FUNCTION_BLOCK "LKinCtrl_MC_MovePath"   // FB35000, SCL
TITLE = LKinCtrl_MovePath
{ S7_Optimized_Access := 'TRUE' }
AUTHOR : tech.team.motioncontrol@siemens.com
FAMILY : LKinCtrl
VERSION : 3.0
// Core function block of LKinCtrl library:
// executes path motion provided by PathData command list
   VAR_INPUT
      execute : Bool;   // rising edge starts action once
      stop : Bool;   // abort path motion
      interrupt : Bool;   // interrupt path motion
      reset : Bool;   // reset FB / acknowledge errors
      sequenceMode : Int;   // activate sequence mode (0) / single step mode (1)
      pathTransition : DInt;   // initial transition configuration for new path motion (1: use bufferMode and transitionParameter)
      bufferMode : DInt := 1;   // inital bufferMode for new path motion
      transitionParameter : Array[1..5] of LReal;   // initial transitionParameter for new path motion
      configuration : "LKinCtrl_typeConfiguration";   // configuration structure
   END_VAR
   VAR_OUTPUT
      done : Bool;   // TRUE: Commanded functionality has been completed successfully
      busy : Bool;   // TRUE: FB is not finished and new output values can be expected
      active : Bool;   // FB in control of axesGroup / kinematic in motion
      commandAborted : Bool;   // TRUE: Commanded functionality has been aborted by another command
      error : Bool;   // TRUE: An error occurred during the execution of the FB
      status : Word;   // status of the FB
      diagnostics : "LKinCtrl_typeMovePathDiagnostics";   // diagnostics information of FB
      activePathData : String["LKINCTRL_LENGTH_OF_PATHDATA_NAME"];   // name of actual PathData
      activeCmdNo : DInt := 0;   // number of actual PathData set
      remainingDistanceActCmd : LReal;   // remaining distance of actual PathData set
      readyForNextPath : Bool := true;   // TRUE: Next PathData can be triggered
   END_VAR
   VAR_IN_OUT
      axesGroup : TO_Kinematics;   // reference to the axesGroup
      pathData : Variant;   // reference to the PathData
      flags : Array[0.."LKINCTRL_NO_OF_LAST_SETFLAG"] of Bool;   // boolean defined by setFlags in PathCommand
      valueFlags : Array[0.."LKINCTRL_NO_OF_LAST_VALUEFLAG"] of LReal;   // value defined by valueFlags in PathCommand
   END_VAR
   VAR
      statExecuteOld : Bool;   // old value of 'execute' input for edge detection
      statStopOld : Bool;   // old value of 'stop' input for edge detection
      statInterruptOld : Bool;   // old value of 'interrupt' input for edge detection
      statResetOld : Bool;   // old value of 'reset' input for edge detection
      statDone : Bool;   // static value for output 'done'
      statBusy : Bool;   // static value for output 'busy'
      statCommandAborted : Bool;   // static value for output 'commandAborted'
      statError : Bool;   // static value for output 'error'
      statErrorID : Word;   // flagWord for FB output: errorID
      statStatus : Word := 16#7000;   // static value for output 'status'
      statSubfunctionStatus : Word;   // status or return value of called FBs, FCs and system blocks
      statStateExecution : DInt := 0;   // state in the state machine of the FB
      statStatePreBuffering : DInt := 0;   // state in the state machine of the FB
      statDebugState : Bool;   // static variable to debug IF state machine if needed
      statEmptyDiagnostics : "LKinCtrl_typeMovePathDiagnostics";   // empty diagnostics information (for initialization purposes only)
      instLKinCtrl_MC_ExecuteKinMotionCmd : "LKinCtrl_MC_ExecuteKinMotionCmd";
      instLKinCtrl_PreBuffer : "LKinCtrl_PreBuffer";
      statPathDataPreBuffered : "LKinCtrl_typePathData_PreBuf";   // preBuffered PathData elements (internal buffer of path motion commands)
      statPathDataElementPreBuffered : "LKinCtrl_typePathDataElement_PreBuf";   // PathData element to be executed by FB_ExecutePathMotion
      statFlagsBuffer : Struct   // buffer to store flag information for past and actual commands
         writeBufferElement : Int := 1;   // pointer on entry to be written
         bufferElement : Array[1.."LKINCTRL_NO_OF_SETFLAGS_BUFFER_ELEMENTS"] of Struct   // flag information for one specific command (see cmdId)
            pathDataName : String["LKINCTRL_LENGTH_OF_PATHDATA_NAME"];   // PathData name of specific command
            pathDataIdentifier : DInt;   // PathData identifier counter of specific command
            cmdId : DInt;   // cmdId of command in PathData
            isIntermediateCmd : Bool;   // TRUE: command is intermediate command
            setFlags : Array[1.."LKINCTRL_NO_OF_CMD_SETFLAGS"] of "LKinCtrl_typeSetFlagElement_Bool";   // setFlags structure equal to PathData command entry
            valueFlags : Array[1.."LKINCTRL_NO_OF_CMD_VALUEFLAGS"] of "LKinCtrl_typeSetFlagElement_LReal";   // setFlags structure equal to PathData command entry
         END_STRUCT;
      END_STRUCT;
      statLastCmdIdPathdata : DInt;   // static value to store last detected cmd in PathData
      statPathDataPreBufferAddPointerOld : Int;   // old value of 'addPointer' in PathDataPreBuffer
      statReadyForNextPath : Bool := true;   // static value for output 'readyForNextPath'
      statStoreInterruptStateExecution : DInt;   // static store variable for state machine status on interrupt
      statExecutionWaitSingleStep : Bool;   // static bit to wait for execution due to sequenceMode
      statExecutionWaitTimerRunning : Bool;   // static bit to wait for execution due to wait time running
      statWaitMain : Bool;   // static bit to wait for execution due to wait flags
      statWaitValueMain : Bool;   // static bit to wait for execution due to wait value flags
      statPreBufferCmdCtr : Int;   // static counter to run FB LKinCtrl_PreBuffer multiple times
      statWaitFlags : Struct   // static struct to store wait flag information
         waitCtr : Int;   // counter for number of wait flags in one command
         waitFlag : Array[1.."LKINCTRL_NO_OF_CMD_SETFLAGS"] of Int;   // flag number as identifier for flag active as wait flag
      END_STRUCT;
      statWaitValueFlags : Struct   // static struct to store wait valueFlag information
         waitCtr : Int;   // counter for number of wait flags in one command
         waitFlag : Array[1.."LKINCTRL_NO_OF_CMD_VALUEFLAGS"] of Int;   // flag number as identifier for flag active as wait valueFlag
      END_STRUCT;
      statPreBufferedPathDataNameOld : String["LKINCTRL_LENGTH_OF_PATHDATA_NAME"];   // static to store old PathDataName in PathDataPreBuffered
      statPathDataIdentifier : USInt;   // static to identify PathDatas independent of given name
      statPreBufferedCmdIdOld : DInt;   // static to store old cmdId value from PathDataPreBuffered
      statSetFlagsBufferWriteBufferElement_old : Int;   // static to store old setFlagsBuffer write element pointer value
      statExecuterWasDone : Bool;   // static to store done output of executer in case of wait flags at end of path
      statWrittenActiveCmdNo : DInt;   // static to store the last written active command number
      statInterruptedAtStart : Bool;   // static to store if interrupt was executed at start of path
      statInitPos : Array[1..4] of LReal;   // static to store the initial position of the TCP
      statOCSFrames : Array[1..3] of "LKinCtrl_typeFrame";   // static to store the OCS frames from TO_Kinematics
      instLKinCtrl_SetFlagCtrl : "LKinCtrl_SetFlagCtrl";
      instLKinCtrl_ValueFlagCtrl : "LKinCtrl_ValueFlagCtrl";
   END_VAR
   VAR_TEMP
      tempExecute : Bool;   // Temporary value for input 'execute'
      tempStop : Bool;   // Temporary value for input 'stop'
      tempInterrupt : Bool;   // Temporary value for input 'interrupt'
      tempReset : Bool;   // Temporary value for input 'stop'
      tempSequenceMode : Int;   // Temporary value for input 'sequenceMode'
      tempEmptyPathDataElementPreBuffered : "LKinCtrl_typePathDataElement_PreBuf";   // Temporary value for empty pre buffer element
      tempCmdCtr : Int;   // Temporary command counter
      tempFlagsBufferElementCtr : Int;   // Temporary flag buffer counter
      tempPreBufferCallCtr : Int;   // Temporary flag buffer call counter
      tempFlagCmdCounter : Int;   // Temporary flag command counter
      tempFlagResetCmdCounter : Int;   // Temporary flag reset counter
   END_VAR
   VAR CONSTANT
      EX_NO_PROCESSING : Int := 0;   // state machine constant
      EX_RESETTING : Int := 5;   // state machine constant
      EX_INTERRUPT_AT_START : Int := 10;   // state machine constant
      EX_GET_CMD : Int := 30;   // state machine constant
      EX_TRIGGERING_CMD : Int := 50;   // state machine constant
      EX_TRIGGERED_CMD : Int := 55;   // state machine constant
      EX_INTERRUPTING : Int := 70;   // state machine constant
      EX_INTERRUPTED : Int := 75;   // state machine constant
      EX_CONTINUEING : Int := 77;   // state machine constant
      EX_CONTINUED : Int := 78;   // state machine constant
      EX_STOPPING : Int := 80;   // state machine constant
      EX_STOPPED_STATE : Int := 85;   // state machine constant
      EX_ERROR_STATE : Int := 90;   // state machine constant
      EX_ALL_TRIGGERED : Int := 100;   // state machine constant
      PB_NO_PROCESSING : Int := 0;   // state machine constant
      PB_ENABLED : Int := 10;   // state machine constant
      PB_OFF_COMP : Int := 15;   // state machine constant
      PB_DISABLED : Int := 20;   // state machine constant
      STATUS_EXECUTION_FINISHED : Word := 16#0000;   // status execution finished without errors
      STATUS_NO_CALL : Word := 16#7000;   // status no job being currently processed
      STATUS_FIRST_CALL : Word := 16#7001;   // status first call after incoming new job (rising edge 'execute')
      STATUS_SUBSEQUENT_CALL : Word := 16#7002;   // status subsequent call during active processing without further details
      STATUS_FB_RESETTING : Word := 16#7010;   // status FB resetting
      STATUS_WAITING_FOR_PREBUFFERED_CMD : Word := 16#7070;   // status waiting for new command in PathData_Prebuffered
      STATUS_PREBUFFERED_FULL : Word := 16#7071;   // status internal cmd buffer filled completely
      STATUS_CMD_LIN_ACTIVE : Word := 16#7301;   // status linear motion command active at axesgroup
      STATUS_CMD_CIRC_ACTIVE : Word := 16#7302;   // status circular motion command active at axesgroup
      STATUS_PATHMOTION_INTERRUPTED : Word := 16#7303;   // status path motion interrupted
      STATUS_PATHMOTION_STOPPING : Word := 16#7304;   // status path motion stopping
      STATUS_READYFORNEXTPATH : Word := 16#7305;   // status FB ready for next path execution
      STATUS_PATHMOTION_RUNNING : Word := 16#7306;   // status path motion running
      STATUS_EXECUTION_WAITING : Word := 16#7307;   // status path execution waiting due to wait flag, wait time or single step mode
      STATUS_CMD_MOVE_DIRECT_ACTIVE : Word := 16#7308;   // status move direct motion command active at axesgroup
      STATUS_STOP_DUE_TO_ERROR : Word := 16#7309;   // status kinematics is stopped due to an error in FB Executer
      STATUS_COMMAND_ABORTED : Word := 16#7FFF;   // status commanded functionality has been aborted by another command
      ERR_UNDEFINED_STATE : Word := 16#8600;   // error due to an undefined state in state machine
      ERR_EXECUTE_KINMOTIONCMD : Word := 16#8201;   // error due to error in FB LKinCtrl_ExecuteKinMotionCmd
      ERR_WRONG_SEQUENCEMODE : Word := 16#8203;   // error due to invalid sequenceMode on input
      ERR_PATHDATA_PARAMETERS : Word := 16#8204;   // error due to malconfiguration in motion command parameters
      ERR_OFFSET_CALCULATION : Word := 16#8205;   // error due to calculation error in offset compensation
      ERR_ERROR_STILL_PENDING : Word := 16#8207;   // error due to previous not acknowledged error (reset MovePath to acknowledge)
      ERR_SET_FLAG_CONTROL : Word := 16#8208;   // error due to error in set flag control FB
      ERR_VALUE_FLAG_CONTROL : Word := 16#8209;   // error due to error in value flag control FB
      INTERRUPT_AT_START : Bool := FALSE;   // interrupt at start of new path to preload commands
      NO_OF_COMMANDS_PRELOADING : USInt := 3;   // number of commands to be preloaded
   END_VAR
   // transitionParameter[1] := -1.0;
   // statFlagsBuffer.bufferElement[1].cmdId := 0;
   // statFlagsBuffer.bufferElement[1].pathDataName := '';
BEGIN
   //==========================================================================================
   // SIEMENS AG
   // (c)Copyright 2020 All Rights Reserved
   //------------------------------------------------------------------------------------------
   // Library: LKinCtrl
   // Tested with: S7-1517T-3 PN/DP
   // Engineering: TIA Portal V16
   // Restrictions: ---
   // Requirements: S7-1500T FW 2.8
   // Functionality: LKinCtrl_MC_MovePath
   // The FB is executing a sequence to drive a path defined by the user in form of a
   // command list of points and motion commands.
   // 
   // Support: tech.team.motioncontrol@siemens.com
   // Note: Parameter comments are only available in language 'English (United States)'
   //------------------------------------------------------------------------------------------
   // Change log table:
   // Version    Date          Expert in charge    Changes applied
   // 01.00.00   06.02.2018    JR                  First release version v1.0
   // 02.00.00   18.04.2019    JR / FR             V2.0
   // 02.01.00   28.05.2019    JR / FR             V2.1 for LKinLang
   // 02.02.00   28.01.2020    JR / FR             V2.2: Added valueFlags and flagOnlyCmd 
   // 02.02.01   07.02.2020    FR / DF             V2.2.1: Disable Prebuffer when MovePath is stopping/reseting/(done)
   // 02.02.02   12.02.2020    FR                  Fix for loops using wrong flag constant
   // 02.03.00   18.03.2020    FR                  Rework Flag FBs; Fix for interrupt/continue
   // 02.04.00   25.03.2020    FR                  Added preprocessing stop for LKinLang
   // 02.04.01   07.05.2020    FR                  Fix 360° circle with circMode 3
   // 02.04.02   16.07.2020    FR                  Several bugfixes
   // 03.00.00   04.08.2020    FR                  Added MoveDirect and ConveyorTracking; V16/FW2.8.2 required!
   // 03.00.01   06.08.2020    FR                  Bugfix
   // 03.00.02   19.10.2020    FR                  Updated ContourOffset; Updated FlagControl; Bugfixes
   // 03.00.03   23.11.2020    FR                  Updated ContourOffset; Fix in MC_ExecuteKinMotionCmd
   // 03.00.05   01.06.2021    FR                  Fixes in FlagCtrl FBs
   // 03.00.06   06.07.2021    FR                  Updated ContourOffset; Fix in MC_ExecuteKinMotionCmd; Fix in FlagCtrl FBs
   //===========================================================================================

   // Work with temporary value / create process image
   #tempExecute := #execute;
   #tempStop := #stop;
   #tempInterrupt := #interrupt;
   #tempReset := #reset;
   #tempSequenceMode := #sequenceMode;

   REGION TRIGGERING
       //===========================================================================================
       // check for sequenceMode to be activated
       IF #tempSequenceMode = 1 THEN
           // set execution wait bit to stop cmds from being executed (wait in EX_TRIGGERING_CMD)
           #statExecutionWaitSingleStep := TRUE;
           // check for incorrect sequenceMode to be selected
       ELSIF (#tempSequenceMode <> 0 AND #tempSequenceMode <> 1)
           // only check if execution is triggered
           AND #tempExecute = TRUE
       THEN
           // set status accordingly
           #statStatus := #ERR_WRONG_SEQUENCEMODE;
           // set execution state machine
           #statStateExecution := #EX_ERROR_STATE;
       END_IF;

       //===========================================================================================
       // check for rising edge of stop input
       IF (#tempStop = TRUE) AND (#statStopOld = FALSE)
       THEN
           // perform stop procedure
           #statStateExecution := #EX_STOPPING;
           // FR 08.04.2020: Set status and bits here to avoid return when status = STATUS_NO_CALL
           #statStatus := #STATUS_PATHMOTION_STOPPING;
           #statDone := FALSE;
           #statBusy := TRUE;
           #statCommandAborted := FALSE;
           #statError := FALSE;
           #statErrorID := 16#0;


           //===========================================================================================
           // check for rising edge of interrupt input
           // FR 17.03.2020: Added "statDone" to condition
           // FR 09.04.2020: Added stopping status to condition
       ELSIF (#tempInterrupt = TRUE) AND (#statInterruptOld = FALSE) AND (#statDone = FALSE)
           AND #statStatus <> #STATUS_PATHMOTION_STOPPING AND #statStatus <> #STATUS_COMMAND_ABORTED
       THEN
           // FR 11.03.2020: Only save state in some cases
           IF #statStateExecution < #EX_INTERRUPTING
               OR #statStateExecution > #EX_CONTINUED THEN
               // store states of interruption for later continue
               #statStoreInterruptStateExecution := #statStateExecution;
           END_IF;
           // perform interrupt procedure
           #statStateExecution := #EX_INTERRUPTING;
           //===========================================================================================
           // check for rising edge of reset input
       ELSIF (#tempReset = TRUE) AND (#statResetOld = FALSE)
           // interlock reset during execution
           AND (#statBusy = FALSE)
       THEN
           // perform reset procedure
           #statStateExecution := #EX_RESETTING;
           #statStatePreBuffering := #PB_NO_PROCESSING;
           // set status accordingly
           #statStatus := #STATUS_FB_RESETTING;
           //===========================================================================================
           // check for rising edge of execute input
       ELSIF (#tempExecute = TRUE) AND (#statExecuteOld = FALSE)
           AND (#stop = FALSE) AND (#interrupt = FALSE)
       THEN // First call; initialize FB
           #statDone := FALSE;
           #statCommandAborted := FALSE;
           #statError := FALSE;
           #statErrorID := 16#0;

           // ERROR on start
           //===========================================================================================
           // check for state machine to be in error state from previous (not acknowledged) error
           IF #statStateExecution = #EX_ERROR_STATE THEN
             // State machine - do not start cmd execution and wait in error state
             //------------------------------------------------------------------------------------------
             // no changes to PreBuffer state machine
             #statStateExecution := #EX_ERROR_STATE;
             #statStatePreBuffering := #PB_NO_PROCESSING;

             // check for error already detected before execute in this cycle (e.g. wrong sequenceMode / other faulty inputs)
             IF #statStatus = #ERR_WRONG_SEQUENCEMODE THEN
               // reset statBusy to avoid interlock of reset
               #statBusy := FALSE;
             ELSE
               // set status to set error bit
               #statStatus := #ERR_ERROR_STILL_PENDING;
             END_IF;


             // continue motion in SINGLESTEP mode
             //===========================================================================================
             // check for execution to be waiting for new rising edge
           ELSIF #statStateExecution = #EX_TRIGGERING_CMD
             AND #statExecutionWaitSingleStep = TRUE
           THEN
             // set FB state to busy
             #statBusy := TRUE;
             // reset execution wait bit stopping cmds from being executed (wait in EX_TRIGGERING_CMD)
             #statExecutionWaitSingleStep := FALSE;

             // CONTINUE after interrupt
             //===========================================================================================
             // check for path motion to be interrupted
           ELSIF #statStateExecution = #EX_INTERRUPTED THEN
             // State machine - continue path motion and sequence
             //------------------------------------------------------------------------------------------
             // no changes to PreBuffer state machine
             #statStateExecution := #EX_CONTINUEING;

             // no setting of FB state to busy necessary, interrupt does not reset busy

             // RETRIGGER during running path motion
             // ==========================================================================================
             // check for path motion to be running with all previous cmds executed
           ELSIF #statStateExecution = #EX_ALL_TRIGGERED
           THEN
             // set FB state to busy
             #statBusy := TRUE;

             // // reset last cmdId in PathData depending on type of attached PathData
             #statLastCmdIdPathdata := 0;

             // Reset bit to memorize done output of MC_ExecuteKinMotionCmd
             #statExecuterWasDone := FALSE;

             // state machines - reStart processing
             //------------------------------------------------------------------------------------------
             #statStatePreBuffering := #PB_ENABLED;
             #statStateExecution := #EX_GET_CMD;
             //------------------------------------------------------------------------------------------
             // initialize functionality: reset of variables, diagnostics, etc. (only at reTriggering)
             #statReadyForNextPath := FALSE;

             // set status - added JR 2019/04/16
             #statStatus := #STATUS_SUBSEQUENT_CALL;

             // START of path motion (initial)
             //===========================================================================================
             // check for path motion not to be running already
           ELSIF #axesGroup.StatusMotionQueue.NumberOfCommands = 0         // no commands in MotionQueue
             AND #axesGroup.StatusWord.%X12 = TRUE                       // TO Kinematics in constant velocity
             AND #axesGroup.StatusPath.Velocity = 0.0                    // TO Kinematics standing still
             AND (#axesGroup.StatusWord.%X6                              // no motion job in progress
             OR #axesGroup.StatusConveyor[1].TrackingState <> 0          // If kinematics is in tracking then done (.X6) is not set
             OR #axesGroup.StatusConveyor[2].TrackingState <> 0
             OR #axesGroup.StatusConveyor[3].TrackingState <> 0)
             AND #statStatus <> #STATUS_EXECUTION_WAITING                // Added FR 2019.03.28
           THEN
             //------------------------------------------------------------------------------------------
             // initialize functionality: reset of variables, diagnostics, etc. (only at first call, no reTriggering)
             #statStatus := #STATUS_FIRST_CALL;
             // set FB state to busy
             #statBusy := TRUE;
             #diagnostics := #statEmptyDiagnostics;
             #statSubfunctionStatus := 16#0;
             #statPathDataPreBuffered.addPointerRestarted := FALSE;

             // initialize buffer variables
             //------------------------------------------------------------------------------------------
             // delete PathDataPreBuffered
             FOR #tempCmdCtr := 1 TO "LKINCTRL_NO_OF_PATHDATA_PREBUFFER_ELEMENTS" DO
               #statPathDataPreBuffered.commands[#tempCmdCtr] := #tempEmptyPathDataElementPreBuffered;
             END_FOR;
             // reset PathDataPreBuffered retrievePointer
             #statPathDataPreBuffered.retrievePointer := 1;
             // initialize add pointer in PathData_PreBuffered
             #statPathDataPreBuffered.addPointer := 1;
             #statPathDataPreBuffered.pathDataName := '';
             // delete cmd stored for execution
             #statPathDataElementPreBuffered := #tempEmptyPathDataElementPreBuffered;
             // counter variable PreBuffer call cycles
             #statPreBufferCmdCtr := "LKINCTRL_NO_OF_START_EXECUTE_CMDS";

             // Reset bit to memorize done output of MC_ExecuteKinMotionCmd
             #statExecuterWasDone := FALSE;
             // reset storage static for old PathData identification value
             #statPathDataIdentifier := 0;

             // store actual position - in case of path starting with relative cmd for contour offset compensation
             //------------------------------------------------------------------------------------------
             #statInitPos[1] := #axesGroup.Tcp.x;
             #statInitPos[2] := #axesGroup.Tcp.y;
             #statInitPos[3] := #axesGroup.Tcp.z;
             #statInitPos[4] := #axesGroup.Tcp.a;

             // initialize flag handling variables
             //------------------------------------------------------------------------------------------
             // Reset waitFlags struct
             #statWaitFlags.waitCtr := 0;
             FOR #tempFlagResetCmdCounter := 1 TO "LKINCTRL_NO_OF_CMD_SETFLAGS" DO
               #statWaitFlags.waitFlag[#tempFlagResetCmdCounter] := -1;
             END_FOR;

             // Reset waitValueFlag struct
             #statWaitValueFlags.waitCtr := 0;
             FOR #tempFlagResetCmdCounter := 1 TO "LKINCTRL_NO_OF_CMD_VALUEFLAGS" DO
               #statWaitValueFlags.waitFlag[#tempFlagResetCmdCounter] := -1;
             END_FOR;

             // reset setFlagsBuffer variables
             #statFlagsBuffer.writeBufferElement := 1;
             #statSetFlagsBufferWriteBufferElement_old := 1;

             // #reset setFlagBuffer
             FOR #tempFlagsBufferElementCtr := 1 TO "LKINCTRL_NO_OF_SETFLAGS_BUFFER_ELEMENTS" DO
               FOR #tempFlagResetCmdCounter := 1 TO "LKINCTRL_NO_OF_CMD_SETFLAGS" DO
                 #statFlagsBuffer.bufferElement[#tempFlagsBufferElementCtr].setFlags[#tempFlagResetCmdCounter].flag := -1;
                 #statFlagsBuffer.bufferElement[#tempFlagsBufferElementCtr].setFlags[#tempFlagResetCmdCounter].flagMode := 0;
                 #statFlagsBuffer.bufferElement[#tempFlagsBufferElementCtr].setFlags[#tempFlagResetCmdCounter].remainingDistance := 0.0;
               END_FOR;
               FOR #tempFlagResetCmdCounter := 1 TO "LKINCTRL_NO_OF_CMD_VALUEFLAGS" DO
                 #statFlagsBuffer.bufferElement[#tempFlagsBufferElementCtr].valueFlags[#tempFlagResetCmdCounter].flag := -1;
                 #statFlagsBuffer.bufferElement[#tempFlagsBufferElementCtr].valueFlags[#tempFlagResetCmdCounter].flagMode := 0;
                 #statFlagsBuffer.bufferElement[#tempFlagsBufferElementCtr].valueFlags[#tempFlagResetCmdCounter].remainingDistance := 0.0;
                 #statFlagsBuffer.bufferElement[#tempFlagsBufferElementCtr].valueFlags[#tempFlagResetCmdCounter].value := 0.0;
               END_FOR;
               #statFlagsBuffer.bufferElement[#tempFlagsBufferElementCtr].cmdId := 0;
               #statFlagsBuffer.bufferElement[#tempFlagsBufferElementCtr].pathDataName := '';
             END_FOR;

             // Call FBs FlagCtrl for resetting flag handling variables
             #instLKinCtrl_SetFlagCtrl(enable := FALSE,
                                       waitMain => #statWaitMain,
                                       flags := #flags,
                                       waitFlags := #statWaitFlags);

             #instLKinCtrl_ValueFlagCtrl(enable := FALSE,
                                         waitMain => #statWaitValueMain,
                                         valueFlags := #valueFlags,
                                         waitFlags := #statWaitValueFlags);

             // reset other static variables
             //------------------------------------------------------------------------------------------
             #statReadyForNextPath := FALSE;
             #statPathDataPreBuffered.addPointerRestarted := FALSE;
             #statPathDataPreBufferAddPointerOld := 0;
             #statStoreInterruptStateExecution := 0;
             #statWrittenActiveCmdNo := -1;

             // reset last cmdId in PathData depending on type of attached PathData
             #statLastCmdIdPathdata := 0;

             // reset execution wait bit stopping cmds from being executed (wait in EX_TRIGGERING_CMD)for first cmd
             #statExecutionWaitSingleStep := FALSE;
             #statExecutionWaitTimerRunning := FALSE;

             // Reset interrupted flag
             #statInterruptedAtStart := FALSE;

             //------------------------------------------------------------------------------------------
             // call FBs with false
             // FR 11.03.2020: Also reset continueMotion input
             #instLKinCtrl_MC_ExecuteKinMotionCmd(execute := FALSE,
                                                  interrupt := FALSE,
                                                  continueMotion := FALSE,
                                                  reset := FALSE,
                                                  stop := FALSE,
                                                  pathDataElementPreBuf := #statPathDataElementPreBuffered,
                                                  to_Kinematics := #axesGroup);

             #instLKinCtrl_PreBuffer(enable := FALSE,
                                     to_Kinematics := #axesGroup,
                                     pathData := #pathData,
                                     pathDataPreBuf := #statPathDataPreBuffered);
             //------------------------------------------------------------------------------------------

             // state machines - start processing
             //------------------------------------------------------------------------------------------
             #statStatePreBuffering := #PB_ENABLED;
             // Check if interrupt at start is enabled
             IF #INTERRUPT_AT_START = FALSE THEN
               #statStateExecution := #EX_GET_CMD;
             ELSE
               #statStateExecution := #EX_INTERRUPT_AT_START;
             END_IF;
           END_IF;

       ELSIF (#statStatus = #STATUS_FIRST_CALL) THEN
           #statStatus := #STATUS_SUBSEQUENT_CALL;
       END_IF;

       // Edge detection input variables
       #statExecuteOld := #tempExecute;
       #statStopOld := #tempStop;
       #statInterruptOld := #tempInterrupt;
       #statResetOld := #tempReset;

   END_REGION TRIGGERING

   IF (#statStatus = #STATUS_NO_CALL) THEN // Nothing to do -> End here to reduce "system load"
       RETURN;
   END_IF;

   REGION PRE_BUFFERING

       // state reached when no pre buffering is active
       REGION PB_NO_PROCESSING
           IF #statStatePreBuffering = #PB_NO_PROCESSING
               // AND #statDebugState = TRUE
           THEN
               // reset  variable for single step debugging of states
               #statDebugState := FALSE;

               // set enable to false because of reset
               #instLKinCtrl_PreBuffer.enable := FALSE;

               // do nothing
           END_IF;

       END_REGION PB_NO_PROCESSING


       // state reached when  pre buffering is active
       REGION PB_ENABLED
           IF #statStatePreBuffering = #PB_ENABLED
               // AND #statDebugState = TRUE
           THEN
               // reset  variable for single step debugging of states
               #statDebugState := FALSE;

               // set no of calls for PreBuffer
               IF #statStatus <> #STATUS_FIRST_CALL THEN
                   #statPreBufferCmdCtr := "LKINCTRL_NO_OF_SEQ_EXECUTE_CMDS";
               END_IF;

               // FR 14.04.2020: Copy OCS frames from TO_Kinematics
               FOR #tempCmdCtr := 1 TO 3 DO
                   #statOCSFrames[#tempCmdCtr].x := #axesGroup.StatusOcsFrame[#tempCmdCtr].x;
                   #statOCSFrames[#tempCmdCtr].y := #axesGroup.StatusOcsFrame[#tempCmdCtr].y;
                   #statOCSFrames[#tempCmdCtr].z := #axesGroup.StatusOcsFrame[#tempCmdCtr].z;
                   #statOCSFrames[#tempCmdCtr].a := #axesGroup.StatusOcsFrame[#tempCmdCtr].a;
                   #statOCSFrames[#tempCmdCtr].b := #axesGroup.StatusOcsFrame[#tempCmdCtr].b;
                   #statOCSFrames[#tempCmdCtr].c := #axesGroup.StatusOcsFrame[#tempCmdCtr].c;
               END_FOR;

               // enable FB PreBuffer
               #instLKinCtrl_PreBuffer.enable := TRUE;

               // call FB PreBuffer multiple times
               FOR #tempPreBufferCallCtr := 1 TO #statPreBufferCmdCtr DO

                   // rest of state code ==> copy here
                   #instLKinCtrl_PreBuffer(initPathTransition := #pathTransition,
                                           initBufferMode := #bufferMode,
                                           initTransitionParameter := #transitionParameter,
                                           initPos := #statInitPos,
                                           OCSFrames := #statOCSFrames,
                                           configuration := #configuration,
                                           to_Kinematics := #axesGroup,
                                           lastCmdIdPathData => #statLastCmdIdPathdata,
                                           pathData := #pathData,
                                           pathDataPreBuf := #statPathDataPreBuffered);

                   // check for FB PreBuffer to signalize an error
                   IF #instLKinCtrl_PreBuffer.error THEN

                       #statStateExecution := #EX_ERROR_STATE;
                       #statSubfunctionStatus := #instLKinCtrl_PreBuffer.status;
                       //  separate handling for PathData malconfiguration and offset compensation calculation errors
                       IF #statSubfunctionStatus > 16#8300
                           AND #statSubfunctionStatus <= 16#8320
                       THEN
                           // write status information to be error in offset compensation
                           #statStatus := #ERR_OFFSET_CALCULATION;
                       ELSE
                           // write status information to be malparametrization in PathData (no offset compensation)
                           #statStatus := #ERR_PATHDATA_PARAMETERS;
                       END_IF;
                       // exit FOR loop to end pre buffering
                       EXIT;

                   ELSIF #instLKinCtrl_PreBuffer.status = 16#7100 THEN // STATUS_ALL_CMDS_BUFFERED
                       // check for FB PreBuffer to have buffered the last element of the PathData to PathData_PreBuf
                       // go to disable state when PreBuffer is done
                       #statStatePreBuffering := #PB_DISABLED;

                       // exit FOR loop to end pre buffering
                       EXIT;

                   ELSE
                       ; // Do nothing -> Keep buffering
                   END_IF;

               END_FOR;

           END_IF; // End of state PB_ENABLED

       END_REGION PB_ENABLED

       // state reached when pre buffering is active
       REGION PB_DISABLED
           IF #statStatePreBuffering = #PB_DISABLED
               // AND #statDebugState = TRUE
           THEN
               // reset  variable for single step debugging of states
               #statDebugState := FALSE;

               // disable FB PreBuffer after finished execution
               #instLKinCtrl_PreBuffer.enable := FALSE;

               // call FB_PreBuffer with false
               // second call of FB necessary, for PathData with one command only ==> handled in one cycle only
               #instLKinCtrl_PreBuffer(to_Kinematics := #axesGroup,
                                       pathData := #pathData,
                                       pathDataPreBuf := #statPathDataPreBuffered);

           END_IF;
       END_REGION PB_DISABLED



   END_REGION PRE_BUFFERING


   REGION EXECUTION

       // state reached when no processing is active 
       REGION EX_NO_PROCESSING
           IF #statStateExecution = #EX_NO_PROCESSING
               // AND #statDebugState = TRUE
           THEN
               // reset  variable for single step debugging of states
               #statDebugState := FALSE;

               // do nothing and wait for execute trigger

           END_IF;
       END_REGION EX_NO_PROCESSING

       REGION EX_INTERRUPT_AT_START
           IF #statStateExecution = #EX_INTERRUPT_AT_START THEN
               #tempInterrupt := TRUE; // Simulate interrupt input

               IF #instLKinCtrl_MC_ExecuteKinMotionCmd.diagnostics.status = 16#7102 THEN
                   // Interrupted --> Start executing commands
                   #statInterruptedAtStart := TRUE;
                   #statStateExecution := #EX_GET_CMD;
               END_IF;
           END_IF;
       END_REGION EX_INTERRUPT_AT_START


       // state reached when resetting is active 
       REGION EX_RESETTING
           IF #statStateExecution = #EX_RESETTING
               // AND #statDebugState = TRUE
           THEN
               // reset  variable for single step debugging of states
               #statDebugState := FALSE;

               // reset state machines
               //------------------------------------------------------------------------------------------
               #statStateExecution := #EX_NO_PROCESSING;
               #statStatePreBuffering := #PB_NO_PROCESSING;

               // reset store buffer variables
               //------------------------------------------------------------------------------------------
               // delete PathDataPreBuffered
               FOR #tempCmdCtr := 1 TO "LKINCTRL_NO_OF_PATHDATA_PREBUFFER_ELEMENTS" DO
                   #statPathDataPreBuffered.commands[#tempCmdCtr] := #tempEmptyPathDataElementPreBuffered;
               END_FOR;
               // reset PathDataPreBuffered retrievePointer
               #statPathDataPreBuffered.retrievePointer := 1;
               // reset restart bit for PathDataPreBuffered addPointer (also on reEnable in LKinCtrl_PreBuffer)
               #statPathDataPreBuffered.addPointerRestarted := FALSE;
               // addPointer will handled in FB PreBuffer
               #statPathDataPreBuffered.pathDataName := '';
               // delete cmd stored for execution
               #statPathDataElementPreBuffered := #tempEmptyPathDataElementPreBuffered;

               // reset last cmdId in PathData depending on type of attached PathData
               //------------------------------------------------------------------------------------------
               #statLastCmdIdPathdata := 0;

               // Reset bit to memorize done output of MC_ExecuteKinMotionCmd
               #statExecuterWasDone := FALSE;
               // reset storage static for old PathData identification value
               #statPathDataIdentifier := 0;

               // initialize flag handling variables
               //------------------------------------------------------------------------------------------
               // Reset waitFlags struct
               #statWaitFlags.waitCtr := 0;
               FOR #tempFlagResetCmdCounter := 1 TO "LKINCTRL_NO_OF_CMD_SETFLAGS" DO
                   #statWaitFlags.waitFlag[#tempFlagResetCmdCounter] := -1;
               END_FOR;

               // Reset waitValueFlag struct
               #statWaitValueFlags.waitCtr := 0;
               FOR #tempFlagResetCmdCounter := 1 TO "LKINCTRL_NO_OF_CMD_VALUEFLAGS" DO
                   #statWaitValueFlags.waitFlag[#tempFlagResetCmdCounter] := -1;
               END_FOR;

               // reset setFlagsBuffer variables
               #statFlagsBuffer.writeBufferElement := 1;
               #statSetFlagsBufferWriteBufferElement_old := 1;

               // #reset setFlagBuffer
               FOR #tempFlagsBufferElementCtr := 1 TO "LKINCTRL_NO_OF_SETFLAGS_BUFFER_ELEMENTS" DO
                   FOR #tempFlagResetCmdCounter := 1 TO "LKINCTRL_NO_OF_CMD_SETFLAGS" DO
                       #statFlagsBuffer.bufferElement[#tempFlagsBufferElementCtr].setFlags[#tempFlagResetCmdCounter].flag := -1;
                       #statFlagsBuffer.bufferElement[#tempFlagsBufferElementCtr].setFlags[#tempFlagResetCmdCounter].flagMode := 0;
                       #statFlagsBuffer.bufferElement[#tempFlagsBufferElementCtr].setFlags[#tempFlagResetCmdCounter].remainingDistance := 0.0;
                   END_FOR;
                   FOR #tempFlagResetCmdCounter := 1 TO "LKINCTRL_NO_OF_CMD_VALUEFLAGS" DO
                       #statFlagsBuffer.bufferElement[#tempFlagsBufferElementCtr].valueFlags[#tempFlagResetCmdCounter].flag := -1;
                       #statFlagsBuffer.bufferElement[#tempFlagsBufferElementCtr].valueFlags[#tempFlagResetCmdCounter].flagMode := 0;
                       #statFlagsBuffer.bufferElement[#tempFlagsBufferElementCtr].valueFlags[#tempFlagResetCmdCounter].remainingDistance := 0.0;
                       #statFlagsBuffer.bufferElement[#tempFlagsBufferElementCtr].valueFlags[#tempFlagResetCmdCounter].value := 0.0;
                   END_FOR;
                   #statFlagsBuffer.bufferElement[#tempFlagsBufferElementCtr].cmdId := 0;
                   #statFlagsBuffer.bufferElement[#tempFlagsBufferElementCtr].pathDataName := '';
               END_FOR;

               // Call FBs FlagCtrl for resetting flag handling variables
               #instLKinCtrl_SetFlagCtrl(enable := FALSE,
                                         waitMain => #statWaitMain,
                                         flags := #flags,
                                         waitFlags := #statWaitFlags);

               #instLKinCtrl_ValueFlagCtrl(enable := FALSE,
                                           waitMain => #statWaitValueMain,
                                           valueFlags := #valueFlags,
                                           waitFlags := #statWaitValueFlags);

               // reset other static variables
               //------------------------------------------------------------------------------------------
               #statReadyForNextPath := TRUE;//FALSE;
               #statPathDataPreBufferAddPointerOld := 0;
               #statStoreInterruptStateExecution := 0;
               #diagnostics := #statEmptyDiagnostics;
               #statSubfunctionStatus := 16#0;
               #statErrorID := 16#0;
               // reset done bit in case of resetting after completion of path
               #statDone := FALSE;
               // reset cnd aborted bit in case of resetting after stop
               #statCommandAborted := FALSE;

               //------------------------------------------------------------------------------------------
               // call FBs with false
               // FR 11.03.2020: Also reset continueMotion input
               #instLKinCtrl_MC_ExecuteKinMotionCmd(execute := FALSE,
                                                    interrupt := FALSE,
                                                    continueMotion := FALSE,
                                                    reset := TRUE,
                                                    pathDataElementPreBuf := #statPathDataElementPreBuffered,
                                                    to_Kinematics := #axesGroup);


               #instLKinCtrl_PreBuffer(enable := FALSE,
                                       to_Kinematics := #axesGroup,
                                       pathData := #pathData,
                                       pathDataPreBuf := #statPathDataPreBuffered);
               //------------------------------------------------------------------------------------------

               // set status ==> FB will be executed once, next cycle no exection by return
               #statStatus := #STATUS_NO_CALL;

           END_IF;
       END_REGION EX_RESETTING


       // state reached new command should be provided from PathData_PreBuffered to LKinCtrl_ExecuteKinMotionCmd 
       REGION EX_GET_CMD
           IF #statStateExecution = #EX_GET_CMD
               // AND #statDebugState = TRUE
           THEN
               // reset  variable for single step debugging of states
               #statDebugState := FALSE;

               // check for lastCmdIdPathInData to be recognized after last execution of EX_TRIGGERED_CMD
               IF #statPathDataElementPreBuffered.cmdID = #statLastCmdIdPathdata
                   AND #statPathDataElementPreBuffered.isIntermediateCmd = FALSE
               THEN
                   // skip GET_NEW_CMD and go back to EX_TRIGGERED_CMD
                   #statStateExecution := #EX_TRIGGERED_CMD;
               ELSE
                   // provide new single cmd from PathData_PreBuffered according to the pointer status
                   //------------------------------------------------------------------------------------------
                   // FR: Adapted IF condition 2019.03.28
                   // check for retrievePointer not to pass addPointer
                   // check PathDataPreBuf to have empty slots (retrievePointer may not pass addPointer) 
                   IF (#statPathDataPreBuffered.retrievePointer <(* = *)#statPathDataPreBuffered.addPointer AND #statPathDataPreBuffered.addPointerRestarted = FALSE
                       // interlock when 'empty' config cmd is buffered !?
                       AND NOT (#statPathDataPreBuffered.retrievePointer = #statPathDataPreBuffered.addPointer AND #instLKinCtrl_PreBuffer.preBufferLockDueToConfigCmd)
                       // interlock when subsequent cmds are deactivated
                       AND NOT (#statPathDataPreBuffered.retrievePointer = #statPathDataPreBuffered.addPointer AND #instLKinCtrl_PreBuffer.statSubsequentDeactCmdCtr > 0)
                       // interlock as long as bufferLocked
                       (* AND #statPathDataPointers.bufferLocked = FALSE *)) // Handled in PreBuffer FR: 2019.03.28
                       // check for pointer restart asynchronously (addPointer restart before retrievePointer)
                       OR (#statPathDataPreBuffered.addPointerRestarted = TRUE AND #statPathDataPreBuffered.retrievePointer > #statPathDataPreBuffered.addPointer)
                       OR (#statPathDataPreBuffered.addPointerRestarted = TRUE AND #statStatus = #STATUS_FIRST_CALL)
                       // positive condition to run in case of offset compensation
                       OR (#statPathDataPreBuffered.addPointerRestarted = TRUE AND #instLKinCtrl_PreBuffer.preBufferLockDueToConfigCmd)
                   THEN

                       // copy command for execution with FB LKinCtrl_MC_ExecuteKinMotionCmd
                       #statPathDataElementPreBuffered := #statPathDataPreBuffered.commands[#statPathDataPreBuffered.retrievePointer];

                       // PathData identifier number - setting
                       //------------------------------------------------------------------------------------------
                       // detect change of PathData - new cmdId smaller or equal to last one ==> new Path
                       IF #statPathDataElementPreBuffered.cmdID <= #statPreBufferedCmdIdOld
                           OR #statPathDataElementPreBuffered.pathDataName <> #statPreBufferedPathDataNameOld
                       THEN
                           // handle PathData identifier counter
                           IF #statPathDataIdentifier < "LKINCTRL_NO_OF_SETFLAGS_BUFFER_ELEMENTS" THEN
                               // increase PathData counter
                               #statPathDataIdentifier += 1;
                           ELSE
                               // restart PathData identifier counter
                               #statPathDataIdentifier := 1;
                           END_IF;
                       ELSE
                           // do nothing
                           ;
                       END_IF;
                       // write PathData identifier in PatDataElement_preBuffered
                       #statPathDataElementPreBuffered.pathDataIdentifier := #statPathDataIdentifier;